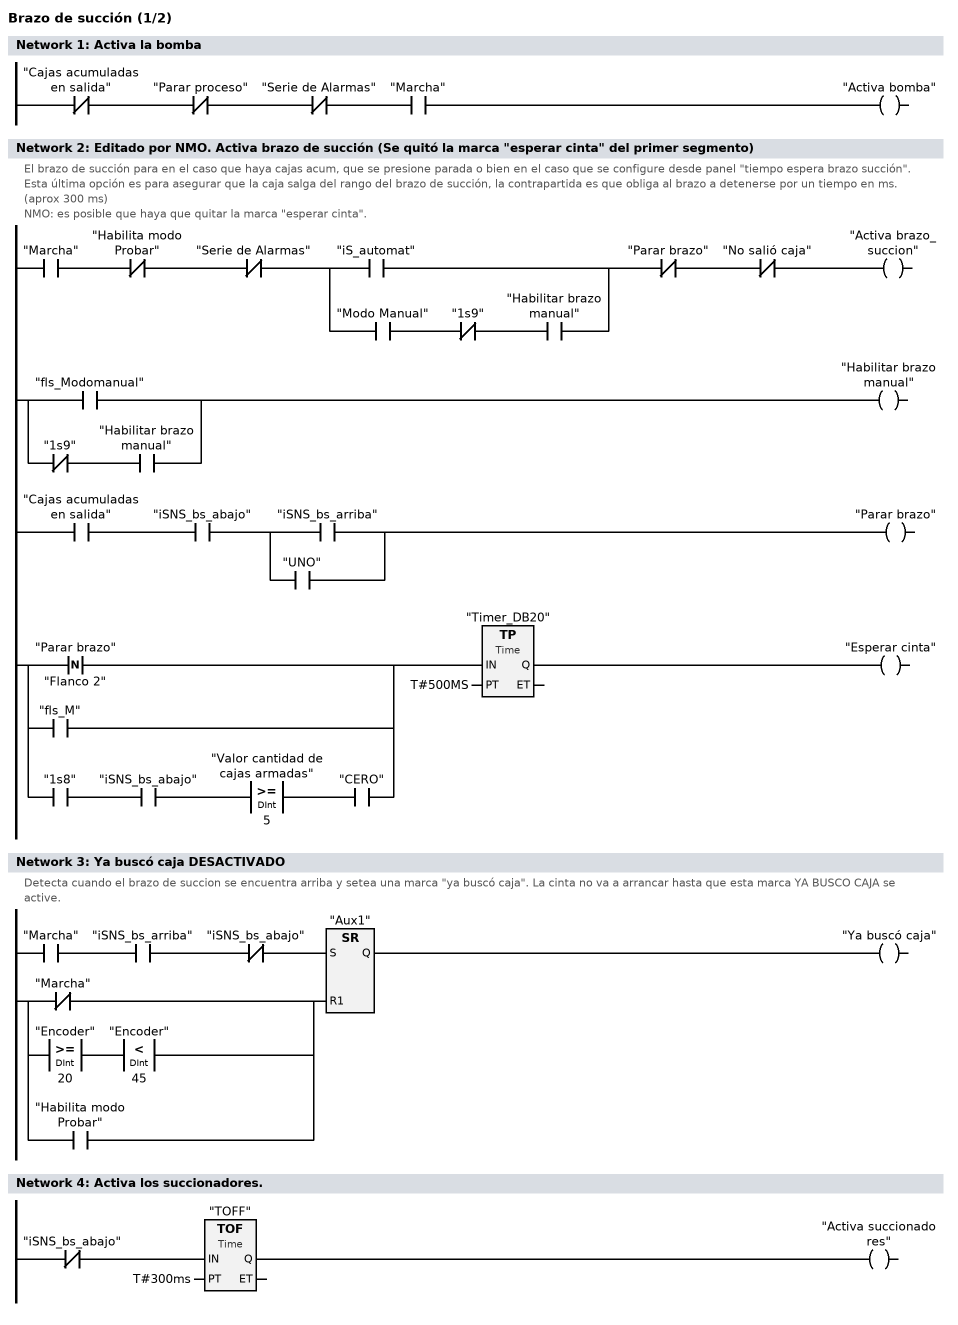
   RUNG wire#powerrail
      I_Contact( "Cajas acumuladas en salida" )
      I_Contact( "Parar proceso" )
      I_Contact( "Serie de Alarmas" )
      Contact( "Marcha" )
      Coil( "Activa bomba" )
   END_RUNG
   // the same network as SCL:
   "Activa bomba" := NOT "Cajas acumuladas en salida" AND NOT "Parar proceso" AND NOT "Serie de Alarmas" AND "Marcha";
END_REGION

REGION Network 2: Editado por NMO. Activa brazo de succión (Se quitó la marca "esperar cinta" del primer segmento)
   // El brazo de succión para en el caso que haya cajas acum, que se presione parada o bien en el caso que se configure desde panel "tiempo espera brazo succión". Esta última opción es para asegurar que la caja salga del rango del brazo de succión, la contrapartida es que obliga al brazo a detenerse por un tiempo en ms. (aprox 300 ms)
   // NMO: es posible que haya que quitar la marca "esperar cinta".
   "Activa brazo_succion" := "Marcha" AND NOT "Habilita modo Probar" AND NOT "Serie de Alarmas" AND ("iS_automat" OR ("Modo Manual" AND NOT "1s9" AND "Habilitar brazo manual")) AND NOT "Parar brazo" AND NOT "No salió caja";
   "Habilitar brazo manual" := "fls_Modomanual" OR (NOT "1s9" AND "Habilitar brazo manual");
   "Parar brazo" := "Cajas acumuladas en salida" AND "iSNS_bs_abajo" AND ("iSNS_bs_arriba" OR "UNO");
   #_w1 := NOT "Parar brazo" AND "Flanco 2";   // falling edge of "Parar brazo"
   "Flanco 2" := "Parar brazo";
   "Timer_DB20".TP(IN := #_w1 OR "fls_M" OR ("1s8" AND "iSNS_bs_abajo" AND ("Valor cantidad de cajas armadas" >= 5) AND "CERO"),
                   PT := T#500MS);
   "Esperar cinta" := "Timer_DB20".Q;
END_REGION

REGION Network 3: Ya buscó caja DESACTIVADO
   // Detecta cuando el brazo de succion se encuentra arriba y setea una marca "ya buscó caja". La cinta no va a arrancar hasta que esta marca YA BUSCO CAJA se active.
   RUNG wire#powerrail
      Contact( "Marcha" )
      Contact( "iSNS_bs_arriba" )
      I_Contact( "iSNS_bs_abajo" )
      S_SR(operand := "Aux1", r1 := wire#w1)
      Coil( "Ya buscó caja" )
   END_RUNG
   RUNG wire#powerrail
      I_Contact( "Marcha" )
   END_RUNG wire#w1
   RUNG wire#powerrail
      { S7_Templates := "SrcType := DInt" } GE_Contact(in1 := "Encoder", in2 := 20)
      { S7_Templates := "SrcType := DInt" } LT_Contact(in1 := "Encoder", in2 := 45)
   END_RUNG wire#w1
   RUNG wire#powerrail
      Contact( "Habilita modo Probar" )
   END_RUNG wire#w1
   // the same network as SCL:
   IF "Marcha" AND "iSNS_bs_arriba" AND NOT "iSNS_bs_abajo" THEN
       "Aux1" := TRUE;   // SR flip-flop
   END_IF;
   IF NOT "Marcha" OR (("Encoder" >= 20) AND ("Encoder" < 45)) OR "Habilita modo Probar" THEN
       "Aux1" := FALSE;
   END_IF;
   "Ya buscó caja" := "Aux1";
END_REGION

REGION Network 4: Activa los succionadores.
   "TOFF".TOF(IN := NOT "iSNS_bs_abajo", PT := T#300ms);
   "Activa succionadores" := "TOFF".Q;
END_REGION

REGION Network 5: Cuando el brazo llega hasta abajo, lo detiene por 300 ms para asegurar que la caja salió de su rango. DESACTIVADO
   // DESACTIVADO
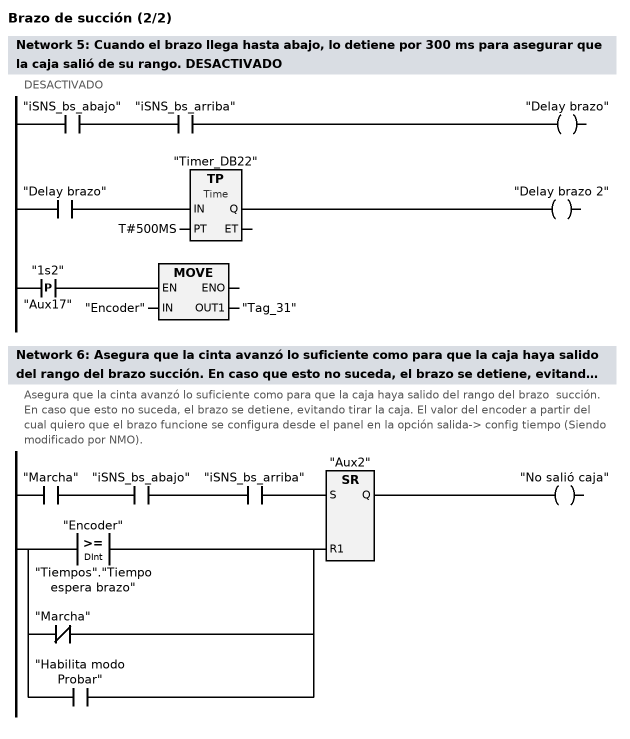
   "Delay brazo" := "iSNS_bs_abajo" AND "iSNS_bs_arriba";
   "Timer_DB22".TP(in := "Delay brazo", pt := T#500MS);
   "Delay brazo 2" := "Timer_DB22".q;
   #_w1 := "1s2" AND NOT "Aux17";   // rising edge of "1s2"
   "Aux17" := "1s2";
   IF #_w1 THEN "Tag_31" := "Encoder"; END_IF;
END_REGION

REGION Network 6: Asegura que la cinta avanzó lo suficiente como para que la caja haya salido del rango del brazo succión. En caso que esto no suceda, el brazo se detiene, evitando tirar la caja
   // Asegura que la cinta avanzó lo suficiente como para que la caja haya salido del rango del brazo  succión. En caso que esto no suceda, el brazo se detiene, evitando tirar la caja. El valor del encoder a partir del cual quiero que el brazo funcione se configura desde el panel en la opción salida-> config tiempo (Siendo modificado por NMO).
   RUNG wire#powerrail
      Contact( "Marcha" )
      Contact( "iSNS_bs_abajo" )
      Contact( "iSNS_bs_arriba" )
      S_SR(operand := "Aux2", r1 := wire#w1)
      Coil( "No salió caja" )
   END_RUNG
   RUNG wire#powerrail
      { S7_Templates := "SrcType := DInt" } GE_Contact(in1 := "Encoder", in2 := "Tiempos"."Tiempo espera brazo")
   END_RUNG wire#w1
   RUNG wire#powerrail
      I_Contact( "Marcha" )
   END_RUNG wire#w1
   RUNG wire#powerrail
      Contact( "Habilita modo Probar" )
   END_RUNG wire#w1
   // the same network as SCL:
   IF "Marcha" AND "iSNS_bs_abajo" AND "iSNS_bs_arriba" THEN
       "Aux2" := TRUE;   // SR flip-flop
   END_IF;
   IF ("Encoder" >= "Tiempos"."Tiempo espera brazo") OR NOT "Marcha" OR "Habilita modo Probar" THEN
       "Aux2" := FALSE;
   END_IF;
   "No salió caja" := "Aux2";
END_REGION
END_FUNCTION

ORGANIZATION_BLOCK "Main"   // OB1, LAD, ProgramCycle
TITLE = "Main Program Sweep (Cycle)"
{ S7_Optimized_Access := 'FALSE' }
VERSION : 0.1
BEGIN

REGION Network 1: Inversión de algunas entradas
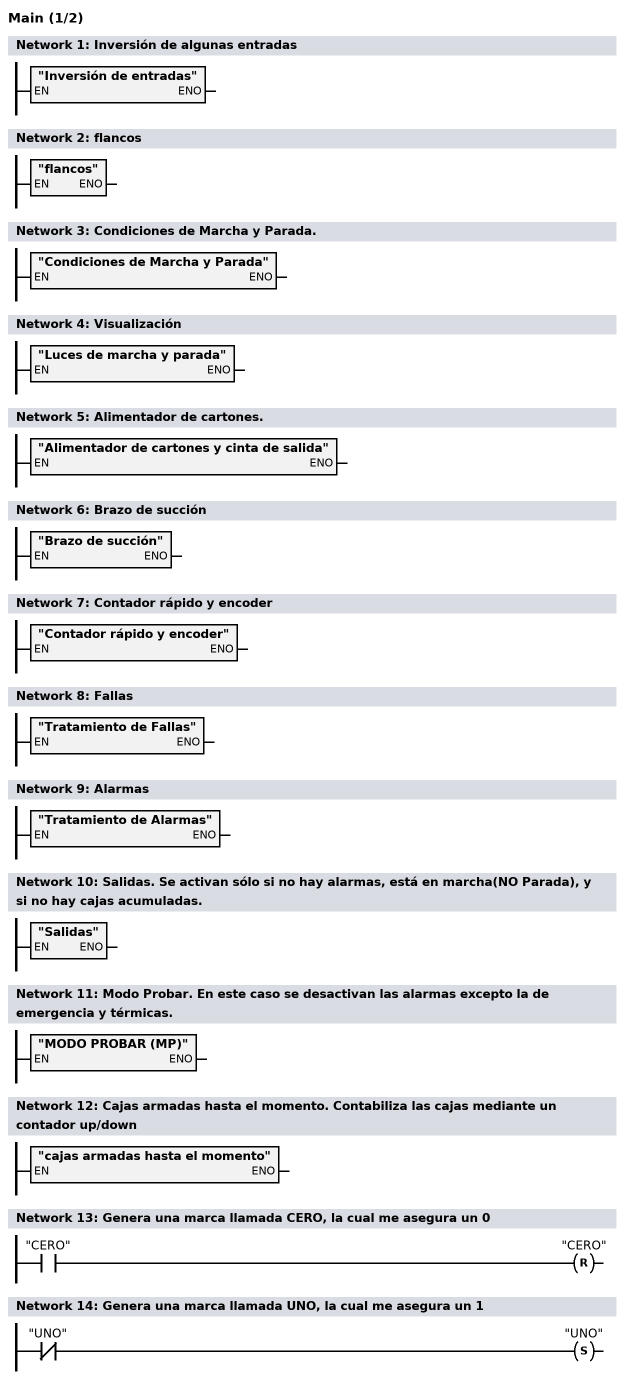
   RUNG wire#powerrail
      "Inversión de entradas"()
   END_RUNG
   // the same network as SCL:
   "Inversión de entradas"();
END_REGION

REGION Network 2: flancos
   RUNG wire#powerrail
      "flancos"()
   END_RUNG
   // the same network as SCL:
   "flancos"();
END_REGION

REGION Network 3: Condiciones de Marcha y Parada.
   RUNG wire#powerrail
      "Condiciones de Marcha y Parada"()
   END_RUNG
   // the same network as SCL:
   "Condiciones de Marcha y Parada"();
END_REGION

REGION Network 4: Visualización
   RUNG wire#powerrail
      "Luces de marcha y parada"()
   END_RUNG
   // the same network as SCL:
   "Luces de marcha y parada"();
END_REGION

REGION Network 5: Alimentador de cartones.
   RUNG wire#powerrail
      "Alimentador de cartones y cinta de salida"()
   END_RUNG
   // the same network as SCL:
   "Alimentador de cartones y cinta de salida"();
END_REGION

REGION Network 6: Brazo de succión
   RUNG wire#powerrail
      "Brazo de succión"()
   END_RUNG
   // the same network as SCL:
   "Brazo de succión"();
END_REGION

REGION Network 7: Contador rápido y encoder
   RUNG wire#powerrail
      "Contador rápido y encoder"()
   END_RUNG
   // the same network as SCL:
   "Contador rápido y encoder"();
END_REGION

REGION Network 8: Fallas
   RUNG wire#powerrail
      "Tratamiento de Fallas"()
   END_RUNG
   // the same network as SCL:
   "Tratamiento de Fallas"();
END_REGION

REGION Network 9: Alarmas
   RUNG wire#powerrail
      "Tratamiento de Alarmas"()
   END_RUNG
   // the same network as SCL:
   "Tratamiento de Alarmas"();
END_REGION

REGION Network 10: Salidas. Se activan sólo si no hay alarmas, está en marcha(NO Parada), y si no hay cajas acumuladas.
   RUNG wire#powerrail
      "Salidas"()
   END_RUNG
   // the same network as SCL:
   "Salidas"();
END_REGION

REGION Network 11: Modo Probar. En este caso se desactivan las alarmas excepto la de emergencia y térmicas.
   RUNG wire#powerrail
      "MODO PROBAR (MP)"()
   END_RUNG
   // the same network as SCL:
   "MODO PROBAR (MP)"();
END_REGION

REGION Network 12: Cajas armadas hasta el momento. Contabiliza las cajas mediante un contador up/down
   RUNG wire#powerrail
      "cajas armadas hasta el momento"()
   END_RUNG
   // the same network as SCL:
   "cajas armadas hasta el momento"();
END_REGION

REGION Network 13: Genera una marca llamada CERO, la cual me asegura un 0
   RUNG wire#powerrail
      Contact( "CERO" )
      R_Coil( "CERO" )
   END_RUNG
   // the same network as SCL:
   IF "CERO" THEN "CERO" := FALSE; END_IF;
END_REGION

REGION Network 14: Genera una marca llamada UNO, la cual me asegura un 1
   RUNG wire#powerrail
      I_Contact( "UNO" )
      S_Coil( "UNO" )
   END_RUNG
   // the same network as SCL:
   IF NOT "UNO" THEN "UNO" := TRUE; END_IF;
END_REGION

REGION Network 15: Secuencia Principal
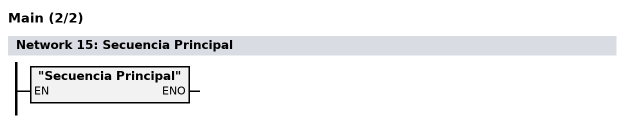
   RUNG wire#powerrail
      "Secuencia Principal"()
   END_RUNG
   // the same network as SCL:
   "Secuencia Principal"();
END_REGION
END_ORGANIZATION_BLOCK

(* ===== HMI "HMI_RT_1" =====
connection "Conexión_HMI": ETHERNET, SMART_S7_1200_OMS

HMI tags "Tabla de variables estándar"
   "Alarmas_1" : Word, 1 s
   "Alarmas_2" : Word, 1 s
   "iAveria-reposicion" : Bool = PLC "iAveria-reposicion", 1 s
   "olmpR" : Bool = PLC "oLmpR", 1 s
   "serie de fallas" : Bool = PLC "Serie de fallas", 1 s
   "Rearme desde panel" : Bool = PLC "Rearme desde panel", 1 s
   "olmpV" : Bool = PLC "oLmpV", 1 s
   "SNS_carton en area de colado" : Bool = PLC "iSNS_carton en area de colado", 1 s
   "SNS_bs_arriba" : Bool = PLC "iSNS_bs_arriba", 1 s
   "SNS_bs_abajo" : Bool = PLC "iSNS_bs_abajo", 1 s
   "sns_nivel_bajo_cartones" : Bool = PLC "iSNS_nivel_bajo_cartones", 1 s
   "SNSpush_atras" : Bool = PLC "iSNSpush_atras", 1 s
   "SNSpush_adel" : Bool = PLC "iSNSpush_adel", 1 s
   "SNSpegamento en depósito" : Bool = PLC "iSNSpegamento en depósito", 1 s
   "SNScaja_trab" : Bool = PLC "iSNScaja_trab", 1 s
   "SNSalp" : Bool = PLC "iSNSalp", 1 s
   "SNScajas_acumuladas" : Bool = PLC "iSnsCajaCerrada", 1 s
   "om_cinta_principal" : Bool = PLC "oM_cinta_principal", 1 s
   "om_bomba" : Bool = PLC "oM_bomba", 1 s
   "oencola" : Bool = PLC "oBoquilla_Encoladora", 1 s
   "om_brazo_succ" : Bool = PLC "oM_brazo_succión", 1 s
   "om_pusher" : Bool = PLC "oM_pusher", 1 s
   "om_cinta_sal" : Bool = PLC "oM_cinta_sal", 1 s
   "osucción" : Bool = PLC "oVálvula_Succión", 1 s
   "oagarra_solapas" : Bool = PLC "oAgarra_solapas", 1 s
   "ocierra_solapa" : Bool = PLC "oCierra_solapa", 1 s
   "opinza" : Bool = PLC "oPinza", 1 s
   "oretB" : Bool = PLC "oRetB", 1 s
   "oretC" : Bool = PLC "oRetC", 1 s
   "oalim_cart" : Bool = PLC "oAlim_cart", 1 s
   "opusher_out" : Bool = PLC "oPusher_out", 1 s
   "iemergencia" : Bool = PLC "iEmergencia", 1 s
   "Emergencia desde panel" : Bool = PLC "Emergencia desde panel", 1 s
   "valor del encoder" : DWord = PLC "Valor del encoder", 100 ms
   "Marcha desde panel" : Bool = PLC "Marcha desde panel", 1 s
   "Parada desde panel" : Bool = PLC "Parada", 1 s
   "S_automat" : Bool = PLC "iS_automat", 1 s
   "S_Probar" : Bool = PLC "iS_Probar", 1 s
   "Modo Manual" : Bool = PLC "Modo Manual", 1 s
   "K_encol_on" : Bool = PLC "iK_encol_on", 1 s
   "Valor cantidad de cajas armadas" : DWord = PLC "Valor cantidad de cajas armadas", 1 s
   "Almacena el valor encolado experimental" : DWord = PLC "Exp Almacena el valor encolado experimental", 1 s
   "ifase0" : Bool = PLC "iFase0", 1 s
   "MPbrazo de succión arriba" : Bool = PLC "MPbrazo de succión arriba", 1 s
   "MPbrazo de succión abajo" : Bool = PLC "MPbrazo de succión abajo", 1 s
   "MPbotón activar pusher" : Bool = PLC "MPbotón activar pusher", 1 s
   "MPbotón Agarra solapas" : Bool = PLC "MPbotón Agarra solapas", 1 s
   "MPbotón activar retenedores de caja" : Bool = PLC "MPbotón activar retenedores de caja", 1 s
   "MPbotón Avanzar cinta por tramos" : Bool = PLC "MPbotón Avanzar cinta por tramos", 1 s
   "MPbotón alimentador de cartones" : Bool = PLC "MPbotón alimentador de cartones", 1 s
   "MPbotón Cierra solapa" : Bool = PLC "MPbotón Cierra solapa", 1 s
   "MPAcomodar brazo de succión" : Bool = PLC "MPAcomodar brazo de succión", 1 s
   "MPActiva bomba de vacío" : Bool = PLC "MPActiva bomba de vacío", 1 s
   "MPbotón Activar encoladora" : Bool = PLC "MPbotón Activar encoladora", 1 s
   "MPbotón Avanzar cinta" : Bool = PLC "MPbotón Avanzar cinta", 1 s
   "MPboton Activar bomba de vacío" : Bool = PLC "MPboton Activar bomba de vacío", 1 s
   "Rearmar" : Bool = PLC "Rearmar", 1 s
   "serie de Alarmas" : Bool = PLC "Serie de Alarmas", 1 s
   "P" : Bool = PLC "iP", 1 s
   "Marcha" : Bool = PLC "Marcha", 1 s
   "marca de prueba fase 0" : Bool = PLC "Exp marca de prueba fase 0", 1 s
   "Cajas acumuladas en salida" : Bool = PLC "Cajas acumuladas en salida", 1 s
   "k_EXT" : Bool = PLC "k_EXT", 1 s
   "ienable" : Bool = PLC "iEnable", 1 s
   "olinea-emergencia" : Bool = PLC "oLinea-emergencia", 1 s
   "opacker" : Bool = PLC "oPacker", 1 s
   "1s1" : Bool = PLC "1s1", 1 s
   "1s2" : Bool = PLC "1s2", 1 s
   "1s3" : Bool = PLC "1s3", 1 s
   "1s4" : Bool = PLC "1s4", 1 s
   "1s5" : Bool = PLC "1s5", 1 s
   "1s6" : Bool = PLC "1s6", 1 s
   "1s7" : Bool = PLC "1s7", 1 s
   "2s1" : Bool = PLC "2s1", 1 s
   "2s2" : Bool = PLC "2s2", 1 s
   "2s3" : Bool = PLC "2s3", 1 s
   "2s4" : Bool = PLC "2s4", 1 s
   "2s5" : Bool = PLC "2s5", 1 s
   "2s6" : Bool = PLC "2s6", 1 s
   "boton activar fingers" : Bool = PLC "Boton activar fingers", 1 s
   "osep_fing" : Bool = PLC "oSep_fing", 1 s
   "botón packer" : Bool = PLC "Botón packer", 1 s
   "oquick_out" : Bool = PLC "oQuick_out", 1 s
   "boton quick out" : Bool = PLC "Boton quick out", 1 s
   "Valor del encoder para calc encolado" : DWord = PLC "Exp valor del encoder para calc encolado", 1 s
   "marca aux id118" : Bool = PLC "Exp marca aux id118", 1 s
   "Pulsador modo manual" : Bool = PLC "Pulsador modo manual", 1 s
   "MPvalor actual del encoder" : DWord = PLC "MPvalor actual del encoder", 1 s
   "Aviso de cinta descalibrada probar" : Bool = PLC "Aviso de cinta descalibrada probar", 1 s
   "1s8" : Bool = PLC "1s8", 1 s
   "1s9" : Bool = PLC "1s9", 1 s
   "SNScaja_acum" : Bool = PLC "iSNScaja_acum", 1 s
   "datos de encolado_selcaja1000/1500" : Bool, 1 s
   "parar proceso" : Bool = PLC "Parar proceso", 1 s
   "MPActivar cilindro pusher" : Bool = PLC "MPActivar cilindro pusher", 1 s
   "MPboton cilindro push" : Bool = PLC "MPboton cilindro push", 1 s
   "datos de encolado_Iniciosol1cj1000" : DInt, 1 s
   "datos de encolado_finsol1cj1000" : DInt, 1 s
   "datos de encolado_Iniciosol2cj1000" : DInt, 1 s
   "datos de encolado_finsol2cj1000" : DInt, 1 s
   "datos de encolado_Iniciosol1cj1500" : DInt, 1 s
   "datos de encolado_finsol1cj1500" : DInt, 1 s
   "datos de encolado_Iniciosol2cj1500" : DInt, 1 s
   "datos de encolado_finsol2cj1500" : DInt, 1 s
   "Resetear cajas armadas" : Bool = PLC "Resetear cajas armadas", 1 s
   "Tiempos_Tiempo cierra sol" : DInt, 1 s
   "Tiempos_Tiempo espera brazo" : DInt, 1 s
   "Valor encoder pusher salida" : DWord = PLC "Valor encoder pusher salida", 1 s
   "Tiempos_tiempo cajas acum" : DInt, 1 s
   "Tag_33" : Bool = PLC "desactivar", 1 s
   "AjusteEncoder_Hab_Pusher" : DInt, 1 s
   "AjusteEncoder_Dhab_Pusher" : DInt, 1 s
   "AjusteEncoder_Reset" : Bool, 1 s
   "AjusteEncoder_Reset_Val" : DInt, 1 s
   "HMI_Hab. Falla caja trab." : Bool = PLC "HMI_Hab. Falla caja trab.", 1 s
   "Hab_Falla_Caja_Caida" : Bool = PLC "HMI_Hab_Falla_Caja_Caida", 1 s

discrete alarms
   1: '', class Alarmas sin acuse, trigger "Alarmas_1" bit 10
   2: '', class Alarmas sin acuse, trigger "Alarmas_1" bit 9
   3: '', class Alarmas sin acuse, trigger "Alarmas_1" bit 8
   4: '', class Alarmas sin acuse, trigger "Alarmas_1" bit 11
   5: '', class Alarmas sin acuse, trigger "Alarmas_1" bit 12
   6: '', class Alarmas sin acuse, trigger "Alarmas_1" bit 13
   7: '', class Alarmas sin acuse, trigger "Alarmas_1" bit 14
   8: '', class Alarmas sin acuse, trigger "Alarmas_1" bit 15
   9: '', class Alarmas sin acuse, trigger "Alarmas_1" bit 0
   10: '', class Alarmas sin acuse, trigger "Alarmas_1" bit 1
   11: '', class Alarmas sin acuse, trigger "Alarmas_1" bit 2
   12: '', class Alarmas sin acuse, trigger "Alarmas_1" bit 3
   13: '', class Alarmas sin acuse, trigger "Alarmas_1" bit 4
   14: '', class Alarmas sin acuse, trigger "Alarmas_1" bit 5
   15: '', class Alarmas sin acuse, trigger "Alarmas_1" bit 6
   16: '', class Alarmas sin acuse, trigger "Alarmas_1" bit 7
   17: '', class Alarmas sin acuse, trigger "Alarmas_2" bit 8
   18: '', class Alarmas sin acuse, trigger "Alarmas_2" bit 9
   19: '', class Alarmas sin acuse, trigger "Alarmas_2" bit 10
   20: '', class Alarmas sin acuse, trigger "Alarmas_2" bit 11
   21: '', class Alarmas sin acuse, trigger "Alarmas_2" bit 12
   22: '', class Alarmas sin acuse, trigger "Alarmas_2" bit 13

text list "Nombre_imagen_lista_texto": 1 ''; 2 ''; 3 ''; 4 ''

screen "Alarmas" 800x480, template "Plantilla_1"
   AlarmView "Visor de avisos_1" at 5,100 size 785x254
   Button "Botón_1" at 12,364 size 780x68
   TextField "Campo de texto_1" at 140,440 size 122x36
   TextField "Campo de texto_9" at 268,440 size 125x36
   TextField "Campo de texto_10" at 398,440 size 122x36
   TextField "Campo de texto_7" at 0,6 size 800x56

screen "Sensores" 800x480, template "Plantilla_1"
   GraphicIOField "PlotLight_Round_G_2" at 418,156 size 42x34
   GraphicIOField "PlotLight_Round_G_1" at 58,154 size 42x34
   GraphicIOField "PlotLight_Round_G_3" at 58,192 size 42x34
   GraphicIOField "PlotLight_Round_G_4" at 58,228 size 42x34
   GraphicIOField "PlotLight_Round_G_5" at 58,266 size 42x34
   GraphicIOField "PlotLight_Round_G_6" at 58,306 size 42x30
   GraphicIOField "PlotLight_Round_G_8" at 418,192 size 42x34
   GraphicIOField "PlotLight_Round_G_9" at 418,228 size 42x34
   TextField "Campo de texto_2" at 475,154 size 200x27
   GraphicIOField "PlotLight_Round_G_10" at 418,264 size 42x34
   TextField "Campo de texto_3" at 115,154 size 197x27
   TextField "Campo de texto_4" at 112,192 size 191x27
   TextField "Campo de texto_5" at 112,230 size 216x27
   TextField "Campo de texto_6" at 112,268 size 179x27
   TextField "Campo de texto_7" at 112,306 size 167x27
   TextField "Campo de texto_9" at 475,192 size 177x27
   TextField "Campo de texto_10" at 475,228 size 179x27
   TextField "Campo de texto_11" at 475,264 size 205x27
   TextField "Campo de texto_1" at 0,6 size 800x56
   TextField "Campo de texto_8" at 140,440 size 122x36
   TextField "Campo de texto_12" at 268,440 size 125x36
   TextField "Campo de texto_13" at 398,440 size 122x36

screen "Salidas" 800x480, template "Plantilla_1"
   GraphicIOField "PlotLight_Round_G_2" at 438,176 size 42x34
   GraphicIOField "PlotLight_Round_G_1" at 438,360 size 42x34
   GraphicIOField "PlotLight_Round_G_3" at 62,140 size 42x34
   GraphicIOField "PlotLight_Round_G_4" at 62,176 size 42x34
   GraphicIOField "PlotLight_Round_G_5" at 62,212 size 42x34
   GraphicIOField "PlotLight_Round_G_6" at 62,252 size 42x30
   GraphicIOField "PlotLight_Round_G_7" at 62,286 size 42x34
   GraphicIOField "PlotLight_Round_G_8" at 62,324 size 42x34
   GraphicIOField "PlotLight_Round_G_9" at 62,360 size 42x34
   TextField "Campo de texto_2" at 498,176 size 166x27
   GraphicIOField "PlotLight_Round_G_10" at 438,140 size 42x34
   TextField "Campo de texto_3" at 498,362 size 121x27
   TextField "Campo de texto_5" at 120,178 size 139x27
   TextField "Campo de texto_6" at 120,214 size 135x27
   TextField "Campo de texto_7" at 120,252 size 151x27
   TextField "Campo de texto_8" at 120,288 size 143x27
   TextField "Campo de texto_9" at 120,326 size 173x27
   TextField "Campo de texto_11" at 495,138 size 120x27
   GraphicIOField "PlotLight_Round_G_11" at 438,324 size 42x34
   TextField "Campo de texto_12" at 498,326 size 122x27
   GraphicIOField "PlotLight_Round_G_12" at 438,212 size 42x34
   TextField "Campo de texto_13" at 498,214 size 122x27
   GraphicIOField "PlotLight_Round_G_13" at 438,250 size 42x34
   TextField "Campo de texto_14" at 498,252 size 144x27
   GraphicIOField "PlotLight_Round_G_14" at 438,286 size 42x34
   TextField "Campo de texto_15" at 498,288 size 153x27
   TextField "Campo de texto_16" at 120,138 size 187x27
   TextField "Campo de texto_10" at 120,362 size 151x27
   TextField "Campo de texto_4" at 140,440 size 122x36
   TextField "Campo de texto_17" at 268,440 size 125x36
   TextField "Campo de texto_18" at 398,440 size 122x36
   TextField "Campo de texto_1" at 0,6 size 800x56

screen "General" 800x480, template "Plantilla_1"
   TextField "Campo de texto_2" at 40,122 size 134x37
   TextField "Campo de texto_5" at 300,122 size 146x37
   TextField "Campo de texto_6" at 325,122 size 85x37
   IOField "Campo ES_1" at 132,386 size 162x30
   IOField "Campo ES_2" at 138,250 size 520x46
   TextField "Campo de texto_1" at 158,212 size 356x35
   Button "Botón_1" at 585,114 size 190x60
   Button "Botón_2" at 320,310 size 132x44
   TextField "Campo de texto_4" at 28,386 size 78x27
   TextField "Campo de texto_7" at 148,440 size 115x36
   TextField "Campo de texto_8" at 268,440 size 112x36
   TextField "Campo de texto_9" at 385,440 size 138x36
   TextField "Campo de texto_3" at 0,6 size 800x56
   TextField "Campo de texto_10" at 40,122 size 117x37
   TextField "Campo de texto_11" at 329,124 size 93x37

Template "Plantilla_1" 800x480
   DateTimeField "Plantilla_Campo de fecha y hora_1" at 512,54 size 195x30
   GraphicView "Plantilla_Visor de gráficos_1" at 20,14 size 162x40
   TextField "Campo de texto_1" at 5,440 size 132x36
   TextField "Campo de texto_3" at 655,440 size 138x36
   TextField "Campo de texto_5" at 525,440 size 125x36
   TextField "Plantilla_Campo de texto_1" at 20,54 size 122x27

screen "Modo Probar" 800x480, template "Plantilla_1"
   Button "Botón_2" at 160,366 size 222x60
   Button "Botón_3" at 422,366 size 222x60
   Button "Botón_5" at 422,302 size 222x60
   Button "Botón_7" at 422,174 size 222x60
   Button "Botón_8" at 160,302 size 222x60
   Button "Botón_11" at 422,238 size 222x60
   Button "Botón_13" at 422,110 size 222x60
   Button "Botón_15" at 160,110 size 222x60
   Button "Botón_16" at 160,174 size 222x60
   IOField "Campo ES_1" at 60,186 size 78x38
   Button "Botón_1" at 160,238 size 222x60
   TextField "Campo de texto_7" at 0,6 size 800x56
   TextField "Campo de texto_1" at 140,440 size 122x36
   TextField "Campo de texto_9" at 268,440 size 125x36
   TextField "Campo de texto_10" at 398,440 size 122x36

screen "Estado Actual" 800x480, template "Plantilla_1"
   TextField "Campo de texto_1" at 95,156 size 163x27
   TextField "Campo de texto_2" at 95,194 size 184x27
   TextField "Campo de texto_3" at 95,232 size 205x27
   TextField "Campo de texto_4" at 95,270 size 206x27
   TextField "Campo de texto_5" at 95,308 size 153x27
   TextField "Campo de texto_6" at 95,346 size 231x27
   TextField "Campo de texto_7" at 470,156 size 215x27
   TextField "Campo de texto_8" at 470,194 size 228x27
   TextField "Campo de texto_9" at 470,232 size 188x27
   GraphicIOField "PlotLight_Round_G_2" at 40,158 size 42x34
   GraphicIOField "PlotLight_Round_G_1" at 40,196 size 42x34
   GraphicIOField "PlotLight_Round_G_3" at 40,234 size 42x34
   GraphicIOField "PlotLight_Round_G_4" at 40,272 size 42x34
   GraphicIOField "PlotLight_Round_G_5" at 40,310 size 42x34
   GraphicIOField "PlotLight_Round_G_6" at 40,348 size 42x34
   GraphicIOField "PlotLight_Round_G_7" at 415,158 size 42x34
   GraphicIOField "PlotLight_Round_G_8" at 415,196 size 42x34
   GraphicIOField "PlotLight_Round_G_9" at 415,234 size 42x34
   TextField "Campo de texto_10" at 0,6 size 800x56
   TextField "Campo de texto_11" at 140,440 size 122x36
   TextField "Campo de texto_12" at 268,440 size 125x36
   TextField "Campo de texto_13" at 398,440 size 122x36

screen "Colero" 800x480, template "Plantilla_1"
   GraphicIOField "PlotLight_Round_G_13" at 65,194 size 42x34
   TextField "Campo de texto_15" at 125,188 size 213x26
   TextField "Campo de texto_3" at 125,240 size 156x26
   GraphicIOField "PlotLight_Round_G_1" at 65,244 size 42x32
   GraphicIOField "PlotLight_Round_G_2" at 65,290 size 42x34
   TextField "Campo de texto_2" at 125,290 size 222x26
   GraphicIOField "PlotLight_Round_G_3" at 65,144 size 42x34
   TextField "Campo de texto_16" at 125,144 size 177x26
   Button "Botón_7" at 502,346 size 232x60
   TextField "Campo de texto_8" at 140,440 size 122x36
   TextField "Campo de texto_9" at 268,440 size 125x36
   TextField "Campo de texto_10" at 398,440 size 122x36
   TextField "Campo de texto_4" at 0,6 size 800x56

screen "Config - 3" 800x480, template "Plantilla_1"
   IOField "Campo ES_1" at 130,272 size 95x30
   IOField "Campo ES_2" at 135,378 size 95x30
   IOField "Campo ES_3" at 258,272 size 95x30
   IOField "Campo ES_4" at 260,380 size 95x30
   TextField "Campo de texto_2" at 135,238 size 53x27
   TextField "Campo de texto_3" at 132,346 size 53x27
   TextField "Campo de texto_4" at 265,236 size 30x27
   TextField "Campo de texto_5" at 265,346 size 30x27
   IOField "Campo ES_5" at 468,274 size 95x30
   IOField "Campo ES_6" at 472,380 size 95x30
   IOField "Campo ES_7" at 590,276 size 95x30
   IOField "Campo ES_8" at 592,382 size 95x30
   TextField "Campo de texto_7" at 472,236 size 53x27
   TextField "Campo de texto_8" at 470,346 size 53x27
   TextField "Campo de texto_9" at 598,236 size 30x27
   TextField "Campo de texto_10" at 598,346 size 30x27
   TextField "Campo de texto_11" at 170,158 size 129x31
   TextField "Campo de texto_12" at 480,154 size 160x31
   TextField "Campo de texto_14" at 0,6 size 800x56
   TextField "Campo de texto_1" at 135,204 size 82x27
   TextField "Campo de texto_6" at 132,312 size 82x27
   TextField "Campo de texto_13" at 475,204 size 82x27
   TextField "Campo de texto_15" at 472,312 size 82x27
   Switch "Interruptor_1" at 98,106 size 622x46
   TextField "Campo de texto_16" at 140,440 size 122x36
   TextField "Campo de texto_17" at 268,440 size 125x36
   TextField "Campo de texto_18" at 398,440 size 122x36

screen "Config - 1" 800x480, template "Plantilla_1"
   IOField "Campo ES_1" at 272,124 size 85x30
   TextField "Campo de texto_1" at 32,120 size 181x27
   TextField "Campo de texto_2" at 32,286 size 441x27
   IOField "Campo ES_2" at 40,334 size 92x32
   TextField "Campo de texto_3" at 158,320 size 393x52
   TextField "Campo de texto_5" at 32,382 size 492x27
   TextField "Campo de texto_4" at 35,160 size 366x77
   TextField "Campo de texto_7" at 0,6 size 800x56
   TextField "Campo de texto_8" at 140,440 size 122x36
   TextField "Campo de texto_9" at 268,440 size 125x36
   TextField "Campo de texto_10" at 398,440 size 122x36

screen "Config - 2" 800x480, template "Plantilla_1"
   IOField "Campo ES_3" at 242,304 size 180x30
   TextField "Campo de texto_7" at 68,254 size 170x27
   IOField "Campo ES_4" at 242,344 size 180x30
   TextField "Campo de texto_8" at 48,340 size 142x27
   IOField "Campo ES_2" at 70,136 size 165x38
   TextField "Campo de texto_2" at 68,100 size 188x27
   Button "Botón_1" at 250,134 size 150x44
   TextField "Campo de texto_14" at 0,6 size 800x56
   TextField "Campo de texto_1" at 90,302 size 110x27
   IOField "Campo ES_1" at 235,186 size 162x30
   TextField "Campo de texto_4" at 130,186 size 78x27
   TextField "Campo de texto_3" at 140,440 size 122x36
   TextField "Campo de texto_9" at 268,440 size 125x36
   TextField "Campo de texto_10" at 398,440 size 122x36
   Switch "Interruptor_1" at 565,322 size 160x64
   TextField "Campo de texto_5" at 532,258 size 173x52
   Switch "Interruptor_2" at 565,178 size 160x64
   TextField "Campo de texto_6" at 525,116 size 173x52
*)